FUNCTION "LKinLang_TokenizeSlot" : DWord   // FC35483, SCL
TITLE = LKinLang_TokenizeSlot
{ S7_Optimized_Access := 'TRUE' }
AUTHOR : tech.team.motioncontrol@siemens.com
FAMILY : LKinLang
VERSION : 1.1
// The FC separates a slot / line from line buffer in separate tokens
   VAR_INPUT
      lineNumber : UDInt;   // Line number input
      line : String;   // Line content input
      lastIndexOfMerger : Int;   // Last index of merger array
   END_VAR
   VAR_OUTPUT
      tokenizedLine : "LKinLang_typeLineTokens";   // Result of tokenization
   END_VAR
   VAR_IN_OUT
      separators : Array[1.."LKINLANG_NUMBER_OF_SEPARATORS"] of Byte;   // Array of separators
      mergers : Array[1.."LKINLANG_NUMBER_OF_MERGERS"] of Byte;   // Array of mergers
      preprocessorConfig : "LKinLang_typePreProcessorReplacement";   // Configuration structure for preProcessor (search/replace)
      errorString : String;   // Error in string format
   END_VAR
   VAR_TEMP
      tempAsciiLine : String["LKINLANG_LENGTH_OF_ASCII_LINE_STRING"];   // Temporary variable for the string line
      tempSeparatorIndex : DInt;   // Temporary variable for found separator index
      tempAsciiLineLength : Int;   // Temporary variable for the length of the string
      tempSignIndex : Int;   // Temporary counter in the string
      tempSignIndexOld : Int;   // Temporary old value of the counter in the string
      tempTokenIndex : Int;   // Temporary token counter for one line
      tempTypeOfChar : Array[0.."LKINLANG_LENGTH_OF_ASCII_LINE_STRING"] of USInt;   // Type of char in string: 0 = Defauflt; 1=Letter, 2=Number, 3=Merger
      tempTokenizedSlotEmpty : "LKinLang_typeLineTokens";   // Empty structure to delete last result
   END_VAR
   // Ret_Val : Return value of function
   VAR CONSTANT
      ERR_INVALID_LINE_NUMBER : DWord := 16#8200;   // Error due to wrong line number
      ERR_TOKEN_OVERFLOW : DWord := 16#8201;   // Error due to token being too long
      ERR_LINE_TOKEN_OUT_OF_BOUNDS : DWord := 16#8202;   // Error due to counter out of array bounds
   END_VAR
BEGIN
   //==========================================================================================
   // SIEMENS AG
   // (c)Copyright 2019 All Rights Reserved
   //------------------------------------------------------------------------------------------
   // Library: LKinLang
   // Tested with: S7-1517T-3 PN/DP
   // Engineering: TIA Portal V15
   // Restrictions: ---
   // Requirements: S7-1500T FW 2.5
   // Functionality: LKinLang_TokenizeSlot
   // The FC separates a slot / line from line buffer in separate tokens
   // 
   // Support: tech.team.motioncontrol@siemens.com
   // Note: Parameter comments are only available in language 'English (United States)'
   //------------------------------------------------------------------------------------------
   // Change log table:
   // Version    Date          Expert in charge    Changes applied
   // 01.00.00   28.05.2019    FR                  First created version
   // 02.00.00   20.03.2020    FR                  Changed funtion to work with one line only
   //=============================================================================

   // Intitialize values
   #LKinLang_TokenizeSlot := 0;
   #tempTokenIndex := 1;

   //--------------------------------------------------------------------------
   // All lines of Slot (PROGRAM) 
   // Information string access: first character to last character [1..n]
   // In Version 1.0 only one line of Slot (tempLineIndexMin == tempLineIndexMax)
   //--------------------------------------------------------------------------
   // FOR #tempLineIndex := #tempLineIndexMin TO #tempLineIndexMax DO

     // Init tokenized slot 
   #tokenizedLine := #tempTokenizedSlotEmpty;

     // Local copy OF ascii line
     #tempAsciiLine := #line;

     // Call of Pre Processor replacements
     "LKinLang_PreProcessor"(preprocessorConfig := #preprocessorConfig,
                             programLine := #tempAsciiLine);

     // Line which includes only a comment counts as an empty codeline (no G command)        
     "LKinLang_DeleteComment"(#tempAsciiLine);

     // Replace $T through space
     "LKinLang_ReplaceTapsBySpaces"(#tempAsciiLine);

     // Delete more than one spaces
     "LKinLang_DeleteMoreThanOneSpaceInRow"(#tempAsciiLine);

     // Length of ascii line
     #tempAsciiLineLength := LEN(#tempAsciiLine);

     IF #tempAsciiLineLength > 0 THEN
       // Get Tyoe of character --> write into array of USINT
       // Later check only Array and do not use Functions
       FOR #tempSignIndex := 1 TO #tempAsciiLineLength DO
         IF "LKinLang_CharacterIsLetter"(CHAR_TO_BYTE(#tempAsciiLine[#tempSignIndex])) THEN
           #tempTypeOfChar[#tempSignIndex] := 1;
         ELSIF "LKinLang_CharacterIsNumeric"(#tempAsciiLine[#tempSignIndex]) THEN
           #tempTypeOfChar[#tempSignIndex] := 2;
         ELSIF "LKinLang_CharacterIsMerger"(character := #tempAsciiLine[#tempSignIndex], lastIndexOfMerger := #lastIndexOfMerger, mergers := #mergers) THEN
           #tempTypeOfChar[#tempSignIndex] := 3;
         ELSE
           #tempTypeOfChar[#tempSignIndex] := 0;
         END_IF;
       END_FOR;

       #tempSignIndexOld := #tempAsciiLineLength + 1;

       // all characters of line
       FOR #tempSignIndex := #tempAsciiLineLength TO 1 BY -1 DO

         IF #tempTypeOfChar[#tempSignIndex] = 0 THEN // Only check for separator if not merger or letter or numeric: FR 2019.03.13
           REGION CECK_FOR_SEPARATOR
             //Check for separator
             //--------------------------------------------------------------------------------
             // compare sign with all separators
             FOR #tempSeparatorIndex := 1 TO "LKINLANG_NUMBER_OF_SEPARATORS" DO
               // detect separator
               IF #separators[#tempSeparatorIndex] = #tempAsciiLine[#tempSignIndex] THEN
                 IF #tempAsciiLineLength - #tempSignIndex > 0
                   AND #tempSignIndexOld - (#tempSignIndex + 1) > 0
                 THEN
                   IF #tempSignIndexOld - (#tempSignIndex + 1) <= "LKINLANG_LENGTH_OF_TOKEN_STRING" THEN
                     IF #tempTokenIndex > "LKINLANG_MAX_NUMBER_OF_TOKEN_PER_LINE" THEN
                       ;//Error: Array out of bounds 
                       #LKinLang_TokenizeSlot := #ERR_LINE_TOKEN_OUT_OF_BOUNDS;
                       #errorString := CONCAT(IN1 := #errorString, IN2 := 'Error: Tokenization - Overflow. Increase number of token per line - line: ');
                       #errorString := CONCAT(IN1 := #errorString, IN2 := UDINT_TO_STRING(#lineNumber));
                       RETURN;
                     ELSE
                       #tokenizedLine.lineToken[#tempTokenIndex] := MID(IN := #tempAsciiLine, P := #tempSignIndex + 1, L := #tempSignIndexOld - (#tempSignIndex + 1));
                       #tempTokenIndex := #tempTokenIndex + 1;
                     END_IF;
                   ELSE
                     ; // ERROR: Token overflow
                     #LKinLang_TokenizeSlot := #ERR_TOKEN_OVERFLOW;
                     #errorString := CONCAT(IN1 := #errorString, IN2 := 'Error: Tokenization - Overflow. Increase token length - line: ');
                     #errorString := CONCAT(IN1 := #errorString, IN2 := UDINT_TO_STRING(#lineNumber));
                     RETURN;
                   END_IF;
                 END_IF;

                 IF #tempTokenIndex > "LKINLANG_MAX_NUMBER_OF_TOKEN_PER_LINE" THEN
                   ;//Error: Array out of bounds 
                   #LKinLang_TokenizeSlot := #ERR_LINE_TOKEN_OUT_OF_BOUNDS;
                   #errorString := CONCAT(IN1 := #errorString, IN2 := 'Error: Tokenization - Overflow. Increase number of token per line - line: ');
                   #errorString := CONCAT(IN1 := #errorString, IN2 := UDINT_TO_STRING(#lineNumber));
                   RETURN;
                 ELSE
                   #tokenizedLine.lineToken[#tempTokenIndex] := MID(IN := #tempAsciiLine, P := #tempSignIndex, L := 1);
                   #tempTokenIndex := #tempTokenIndex + 1;
                   #tempSignIndexOld := #tempSignIndex;
                 END_IF;
                 EXIT;
               ELSE
                 ;// no match
               END_IF;
             END_FOR;
           END_REGION
         END_IF;

         REGION CHECK_FOR_LETTER_NUMBER
           //--------------------------------------------------------------------------------
           // Separator: Letter -> Number or Number -> letter
           IF #tempSignIndex >= 2 THEN // only possible if it isn´t the last character
             // Changed FR 2019.03.11: Replaced FC call with array
             IF
               ((#tempTypeOfChar[#tempSignIndex] = 2 AND (#tempTypeOfChar[#tempSignIndex - 1] = 1 OR NOT (#tempTypeOfChar[#tempSignIndex - 1] = 2))) // Number -> Letter 
               OR (#tempTypeOfChar[#tempSignIndex] = 1 AND (#tempTypeOfChar[#tempSignIndex - 1] = 2 OR NOT (#tempTypeOfChar[#tempSignIndex - 1] = 1)))) // Letter -> Number
               AND NOT (#tempTypeOfChar[#tempSignIndex - 1] = 3) // Merger to not separate Tokens
             THEN
               // New token found
               IF (#tempSignIndexOld - #tempSignIndex) <= "LKINLANG_LENGTH_OF_TOKEN_STRING" THEN
                 IF #tempTokenIndex > "LKINLANG_MAX_NUMBER_OF_TOKEN_PER_LINE" THEN
                   ;//Error: Array out of bounds 
                   #LKinLang_TokenizeSlot := #ERR_LINE_TOKEN_OUT_OF_BOUNDS;
                   #errorString := CONCAT(IN1 := #errorString, IN2 := 'Error: Tokenization - Overflow. Increase number of token per line - line: ');
                   #errorString := CONCAT(IN1 := #errorString, IN2 := UDINT_TO_STRING(#lineNumber));
                   RETURN;
                 ELSE
                   #tokenizedLine.lineToken[#tempTokenIndex] := MID(IN := #tempAsciiLine, P := #tempSignIndex, L := #tempSignIndexOld - #tempSignIndex);
                   #tempTokenIndex := #tempTokenIndex + 1;
                   #tempSignIndexOld := #tempSignIndex;
                 END_IF;
               ELSE
                 // ERROR: Token overflow
                 #LKinLang_TokenizeSlot := #ERR_TOKEN_OVERFLOW;
                 #errorString := CONCAT(IN1 := #errorString, IN2 := 'Error: Tokenization - Overflow. Increase token length');
                 RETURN;
               END_IF;
             ELSE
               ; // No change in character type --> check next character
             END_IF;
           END_IF;
           //--------------------------------------------------------------------------------
         END_REGION
       END_FOR;

       // Write number of token to structure
       #tokenizedLine.numberOfToken := INT_TO_UINT(#tempTokenIndex);

       // Last few signs
       IF #tempTokenIndex > "LKINLANG_MAX_NUMBER_OF_TOKEN_PER_LINE" THEN
         ;//Error: Array out of bounds 
         #LKinLang_TokenizeSlot := #ERR_LINE_TOKEN_OUT_OF_BOUNDS;
         #errorString := CONCAT(IN1 := #errorString, IN2 := 'Error: Tokenization - Overflow. Increase number of token per line - line: ');
         #errorString := CONCAT(IN1 := #errorString, IN2 := UDINT_TO_STRING(#lineNumber));
         RETURN;
       ELSE
         #tokenizedLine.lineToken[#tempTokenIndex] := MID(IN := #tempAsciiLine, P := 1, L := #tempSignIndexOld - 1);
       END_IF;
       // set token index for next line
       #tempTokenIndex := 1;
       // Write line number of ASCII file for N
       #tokenizedLine.lineNo := #lineNumber;

     ELSE
       // Empty line 
       #tokenizedLine.numberOfToken := 0;
       #tokenizedLine.lineNo := #lineNumber;
     END_IF;

   // END_FOR; //END: All lines of Slot (PROGRAM)
END_FUNCTION

FUNCTION "LKinLang_UpdateModalData" : Void   // FC35484, SCL
TITLE = LKinLang_UpdateModalData
{ S7_Optimized_Access := 'TRUE' }
AUTHOR : tech.team.motioncontrol@siemens.com
FAMILY : LKinLang
VERSION : 1.1
// The FC updates only modal parameters in a given PathData element
   VAR_IN_OUT
      inputPathData : "LKinLang_typePathDataElement";   // input PathData element to be updated
      updatedPathData : "LKinLang_typePathDataElement";   // updated PathData element
   END_VAR
   VAR_TEMP
      tempCounter : Int;   // temporary counter / temporary counter for empty lines
   END_VAR
BEGIN
   //==========================================================================================
   // SIEMENS AG
   // (c)Copyright 2019 All Rights Reserved
   //------------------------------------------------------------------------------------------
   // Library: LKinLang
   // Tested with: S7-1517T-3 PN/DP
   // Engineering: TIA Portal V15
   // Restrictions: ---
   // Requirements: S7-1500T FW 2.5
   // Functionality: LKinLang_UpdateModalData
   // The FC updates only modal parameters in a given PathData element
   // 
   // Support: tech.team.motioncontrol@siemens.com
   // Note: Parameter comments are only available in language 'English (United States)'
   //------------------------------------------------------------------------------------------
   // Change log table:
   // Version    Date          Expert in charge    Changes applied
   // 01.00.00   28.05.2019    FR                  First created version
   // 01.00.02   29.07.2019    FR                  Removed max negative value condition from IFs
   //=============================================================================

   //======================================================================
   // Copy input to output where input is not default and priority is higher
   //======================================================================  


   REGION UPDATE_ALL
     // Check CmdType
     IF #inputPathData.priority.cmdType > #updatedPathData.priority.cmdType THEN
       #updatedPathData.pathDataElement.cmdType := #inputPathData.pathDataElement.cmdType;
       #updatedPathData.priority.cmdType := #inputPathData.priority.cmdType;
     END_IF;

     // Check Coordinates
     // Update Cartesian positions
     IF  #inputPathData.priority.cmdCoordinates.cartesianPosition.x > #updatedPathData.priority.cmdCoordinates.cartesianPosition.x THEN
       #updatedPathData.pathDataElement.cmdCoordinates.cartesianPosition.x := #inputPathData.pathDataElement.cmdCoordinates.cartesianPosition.x;
       #updatedPathData.priority.cmdCoordinates.cartesianPosition.x := #inputPathData.priority.cmdCoordinates.cartesianPosition.x;
     END_IF;
     IF  #inputPathData.priority.cmdCoordinates.cartesianPosition.y > #updatedPathData.priority.cmdCoordinates.cartesianPosition.y THEN
       #updatedPathData.pathDataElement.cmdCoordinates.cartesianPosition.y := #inputPathData.pathDataElement.cmdCoordinates.cartesianPosition.y;
       #updatedPathData.priority.cmdCoordinates.cartesianPosition.y := #inputPathData.priority.cmdCoordinates.cartesianPosition.y;
     END_IF;
     IF  #inputPathData.priority.cmdCoordinates.cartesianPosition.z > #updatedPathData.priority.cmdCoordinates.cartesianPosition.z THEN
       #updatedPathData.pathDataElement.cmdCoordinates.cartesianPosition.z := #inputPathData.pathDataElement.cmdCoordinates.cartesianPosition.z;
       #updatedPathData.priority.cmdCoordinates.cartesianPosition.z := #inputPathData.priority.cmdCoordinates.cartesianPosition.z;
     END_IF;
     IF #inputPathData.priority.cmdCoordinates.cartesianPosition.a > #updatedPathData.priority.cmdCoordinates.cartesianPosition.a THEN
       #updatedPathData.pathDataElement.cmdCoordinates.cartesianPosition.a := #inputPathData.pathDataElement.cmdCoordinates.cartesianPosition.a;
       #updatedPathData.priority.cmdCoordinates.cartesianPosition.a := #inputPathData.priority.cmdCoordinates.cartesianPosition.a;
     END_IF;

     // Check coord system
     IF #inputPathData.priority.cmdCoordinates.coordSystem > #updatedPathData.priority.cmdCoordinates.coordSystem THEN
       #updatedPathData.pathDataElement.cmdCoordinates.coordSystem := #inputPathData.pathDataElement.cmdCoordinates.coordSystem;
       #updatedPathData.priority.cmdCoordinates.coordSystem := #inputPathData.priority.cmdCoordinates.coordSystem;
     END_IF;

     // Check Parameter
     // Check buffer mode
     IF #inputPathData.priority.cmdParameters.bufferMode > #updatedPathData.priority.cmdParameters.bufferMode THEN
       #updatedPathData.pathDataElement.cmdParameters.bufferMode := #inputPathData.pathDataElement.cmdParameters.bufferMode;
       #updatedPathData.priority.cmdParameters.bufferMode := #inputPathData.priority.cmdParameters.bufferMode;
     END_IF;

     // Check dynamic adaption
     IF #inputPathData.priority.cmdParameters.dynamicAdaption > #updatedPathData.priority.cmdParameters.dynamicAdaption THEN
       #updatedPathData.pathDataElement.cmdParameters.dynamicAdaption := #inputPathData.pathDataElement.cmdParameters.dynamicAdaption;
       #updatedPathData.priority.cmdParameters.dynamicAdaption := #inputPathData.priority.cmdParameters.dynamicAdaption;
     END_IF;

     // Check offsetParaNo
     IF #inputPathData.priority.cmdParameters.offsetParameters.offsetParaNo > #updatedPathData.priority.cmdParameters.offsetParameters.offsetParaNo THEN
       #updatedPathData.pathDataElement.cmdParameters.offsetParameters.offsetParaNo := #inputPathData.pathDataElement.cmdParameters.offsetParameters.offsetParaNo;
       #updatedPathData.priority.cmdParameters.offsetParameters.offsetParaNo := #inputPathData.priority.cmdParameters.offsetParameters.offsetParaNo;
     END_IF;

     // Check main path plane
     IF #inputPathData.priority.cmdParameters.offsetParameters.mainPathPlane > #updatedPathData.priority.cmdParameters.offsetParameters.mainPathPlane THEN
       #updatedPathData.pathDataElement.cmdParameters.offsetParameters.mainPathPlane := #inputPathData.pathDataElement.cmdParameters.offsetParameters.mainPathPlane;
       #updatedPathData.priority.cmdParameters.offsetParameters.mainPathPlane := #inputPathData.priority.cmdParameters.offsetParameters.mainPathPlane;
     END_IF;

     // Check orientation direction
     IF #inputPathData.priority.cmdParameters.orientationDirection > #updatedPathData.priority.cmdParameters.orientationDirection THEN
       #updatedPathData.pathDataElement.cmdParameters.orientationDirection := #inputPathData.pathDataElement.cmdParameters.orientationDirection;
       #updatedPathData.priority.cmdParameters.orientationDirection := #inputPathData.priority.cmdParameters.orientationDirection;
     END_IF;

     // Check transition parameter
     FOR #tempCounter := 1 TO 5 DO
       IF #inputPathData.priority.cmdParameters.transitionParameters[#tempCounter] > #updatedPathData.priority.cmdParameters.transitionParameters[#tempCounter] THEN
         #updatedPathData.pathDataElement.cmdParameters.transitionParameters[#tempCounter] := #inputPathData.pathDataElement.cmdParameters.transitionParameters[#tempCounter];
         #updatedPathData.priority.cmdParameters.transitionParameters[#tempCounter] := #inputPathData.priority.cmdParameters.transitionParameters[#tempCounter];
       END_IF;
     END_FOR;

     // Check circle parameters
     // Arc
     IF #inputPathData.priority.cmdParameters.circleParameters.arc > #updatedPathData.priority.cmdParameters.circleParameters.arc THEN
       #updatedPathData.pathDataElement.cmdParameters.circleParameters.arc := #inputPathData.pathDataElement.cmdParameters.circleParameters.arc;
       #updatedPathData.priority.cmdParameters.circleParameters.arc := #inputPathData.priority.cmdParameters.circleParameters.arc;
     END_IF;

     // Circ plane
     IF #inputPathData.priority.cmdParameters.circleParameters.circlePlane > #updatedPathData.priority.cmdParameters.circleParameters.circlePlane THEN
       #updatedPathData.pathDataElement.cmdParameters.circleParameters.circlePlane := #inputPathData.pathDataElement.cmdParameters.circleParameters.circlePlane;
       #updatedPathData.priority.cmdParameters.circleParameters.circlePlane := #inputPathData.priority.cmdParameters.circleParameters.circlePlane;
     END_IF;

     // Circ mode
     IF #inputPathData.priority.cmdParameters.circleParameters.circMode > #updatedPathData.priority.cmdParameters.circleParameters.circMode THEN
       #updatedPathData.pathDataElement.cmdParameters.circleParameters.circMode := #inputPathData.pathDataElement.cmdParameters.circleParameters.circMode;
       #updatedPathData.priority.cmdParameters.circleParameters.circMode := #inputPathData.priority.cmdParameters.circleParameters.circMode;
     END_IF;

     // path choice 
     IF #inputPathData.priority.cmdParameters.circleParameters.pathChoice > #updatedPathData.priority.cmdParameters.circleParameters.pathChoice THEN
       #updatedPathData.pathDataElement.cmdParameters.circleParameters.pathChoice := #inputPathData.pathDataElement.cmdParameters.circleParameters.pathChoice;
       #updatedPathData.priority.cmdParameters.circleParameters.pathChoice := #inputPathData.priority.cmdParameters.circleParameters.pathChoice;
     END_IF;

     // Radius
     IF #inputPathData.priority.cmdParameters.circleParameters.radius > #updatedPathData.priority.cmdParameters.circleParameters.radius THEN
       #updatedPathData.pathDataElement.cmdParameters.circleParameters.radius := #inputPathData.pathDataElement.cmdParameters.circleParameters.radius;
       #updatedPathData.priority.cmdParameters.circleParameters.radius := #inputPathData.priority.cmdParameters.circleParameters.radius;
     END_IF;

     // Aux point
     FOR #tempCounter := 1 TO 3 DO
       IF #inputPathData.priority.cmdParameters.circleParameters.auxPoint[#tempCounter] > #updatedPathData.priority.cmdParameters.circleParameters.auxPoint[#tempCounter] THEN
         #updatedPathData.pathDataElement.cmdParameters.circleParameters.auxPoint[#tempCounter] := #inputPathData.pathDataElement.cmdParameters.circleParameters.auxPoint[#tempCounter];
         #updatedPathData.priority.cmdParameters.circleParameters.auxPoint[#tempCounter] := #inputPathData.priority.cmdParameters.circleParameters.auxPoint[#tempCounter];
       END_IF;
     END_FOR;


     // Check dynamics
     // Velocity
     IF #inputPathData.priority.cmdParameters.pathDynamics.velocity > #updatedPathData.priority.cmdParameters.pathDynamics.velocity THEN
       #updatedPathData.pathDataElement.cmdParameters.pathDynamics.velocity := #inputPathData.pathDataElement.cmdParameters.pathDynamics.velocity;
       #updatedPathData.priority.cmdParameters.pathDynamics.velocity := #inputPathData.priority.cmdParameters.pathDynamics.velocity;
     END_IF;

     // Accelerration
     IF #inputPathData.priority.cmdParameters.pathDynamics.acceleration > #updatedPathData.priority.cmdParameters.pathDynamics.acceleration THEN
       #updatedPathData.pathDataElement.cmdParameters.pathDynamics.acceleration := #inputPathData.pathDataElement.cmdParameters.pathDynamics.acceleration;
       #updatedPathData.priority.cmdParameters.pathDynamics.acceleration := #inputPathData.priority.cmdParameters.pathDynamics.acceleration;
     END_IF;

     // Deceleration
     IF #inputPathData.priority.cmdParameters.pathDynamics.deceleration > #updatedPathData.priority.cmdParameters.pathDynamics.deceleration THEN
       #updatedPathData.pathDataElement.cmdParameters.pathDynamics.deceleration := #inputPathData.pathDataElement.cmdParameters.pathDynamics.deceleration;
       #updatedPathData.priority.cmdParameters.pathDynamics.deceleration := #inputPathData.priority.cmdParameters.pathDynamics.deceleration;
     END_IF;

     // Jerk
     IF #inputPathData.priority.cmdParameters.pathDynamics.jerk > #updatedPathData.priority.cmdParameters.pathDynamics.jerk THEN
       #updatedPathData.pathDataElement.cmdParameters.pathDynamics.jerk := #inputPathData.pathDataElement.cmdParameters.pathDynamics.jerk;
       #updatedPathData.priority.cmdParameters.pathDynamics.jerk := #inputPathData.priority.cmdParameters.pathDynamics.jerk;
     END_IF;

     // Check flags
     FOR #tempCounter := 1 TO "LKINCTRL_NO_OF_CMD_SETFLAGS" DO
       // Check set flag
       IF #inputPathData.priority.setFlags[#tempCounter].flag > #updatedPathData.priority.setFlags[#tempCounter].flag THEN
         #updatedPathData.pathDataElement.setFlags[#tempCounter].flag := #inputPathData.pathDataElement.setFlags[#tempCounter].flag;
         #updatedPathData.priority.setFlags[#tempCounter].flag := #inputPathData.priority.setFlags[#tempCounter].flag;
       END_IF;

       // Check flag mode
       IF #inputPathData.priority.setFlags[#tempCounter].flagMode > #updatedPathData.priority.setFlags[#tempCounter].flagMode THEN
         #updatedPathData.pathDataElement.setFlags[#tempCounter].flagMode := #inputPathData.pathDataElement.setFlags[#tempCounter].flagMode;
         #updatedPathData.priority.setFlags[#tempCounter].flagMode := #inputPathData.priority.setFlags[#tempCounter].flagMode;
       END_IF;

       // Check flag remaining distance
       IF #inputPathData.priority.setFlags[#tempCounter].flagMode > #updatedPathData.priority.setFlags[#tempCounter].remainingDistance THEN
         #updatedPathData.pathDataElement.setFlags[#tempCounter].remainingDistance := #inputPathData.pathDataElement.setFlags[#tempCounter].remainingDistance;
         #updatedPathData.priority.setFlags[#tempCounter].remainingDistance := #inputPathData.priority.setFlags[#tempCounter].remainingDistance;
       END_IF;
     END_FOR;

     // Check value flags
     FOR #tempCounter := 1 TO "LKINCTRL_NO_OF_CMD_VALUEFLAGS" DO
       // Check set flag
       IF #inputPathData.priority.valueFlags[#tempCounter].flag > #updatedPathData.priority.valueFlags[#tempCounter].flag THEN
         #updatedPathData.pathDataElement.valueFlags[#tempCounter].flag := #inputPathData.pathDataElement.valueFlags[#tempCounter].flag;
         #updatedPathData.priority.valueFlags[#tempCounter].flag := #inputPathData.priority.valueFlags[#tempCounter].flag;
       END_IF;

       // Check flag mode
       IF #inputPathData.priority.valueFlags[#tempCounter].flagMode > #updatedPathData.priority.valueFlags[#tempCounter].flagMode THEN
         #updatedPathData.pathDataElement.valueFlags[#tempCounter].flagMode := #inputPathData.pathDataElement.valueFlags[#tempCounter].flagMode;
         #updatedPathData.priority.valueFlags[#tempCounter].flagMode := #inputPathData.priority.valueFlags[#tempCounter].flagMode;
       END_IF;

       // Check flag remaining distance
       IF #inputPathData.priority.valueFlags[#tempCounter].flagMode > #updatedPathData.priority.valueFlags[#tempCounter].remainingDistance THEN
         #updatedPathData.pathDataElement.valueFlags[#tempCounter].remainingDistance := #inputPathData.pathDataElement.valueFlags[#tempCounter].remainingDistance;
         #updatedPathData.priority.valueFlags[#tempCounter].remainingDistance := #inputPathData.priority.valueFlags[#tempCounter].remainingDistance;
       END_IF;
     END_FOR;
   END_REGION
END_FUNCTION

FUNCTION "LKinLang_GetVariable" : Void   // FC35485, SCL
TITLE = LKinLang_GetVariable
{ S7_Optimized_Access := 'TRUE' }
AUTHOR : tech.team.motioncontrol@siemens.com
FAMILY : LKinLang
VERSION : 1.0
// The FC gets the value of a variable and adds it to a string
   VAR_INPUT
      varIndex : Int;   // Variable index
      varType : Int;   // Variable type
   END_VAR
   VAR_IN_OUT
      localVariables : "LKinLang_typeLocalVariables";   // Variables reference list
      interfaceVariables : "LKinLang_typeInterfaceVariables";   // Key token to find variables
      stringExpression : String;   // String expression
   END_VAR
BEGIN
   //==========================================================================================
   // SIEMENS AG
   // (c)Copyright 2020 All Rights Reserved
   //------------------------------------------------------------------------------------------
   // Library: LKinLang
   // Tested with: S7-1517T-3 PN/DP
   // Engineering: TIA Portal V15
   // Restrictions: ---
   // Requirements: S7-1500T FW 2.5
   // Functionality: LKinLang_IsTokenVariable
   // The FC gets the value of a variable and adds it to a string
   // 
   // Support: tech.team.motioncontrol@siemens.com
   // Note: Parameter comments are only available in language 'English (United States)'
   //------------------------------------------------------------------------------------------
   // Change log table:
   // Version    Date          Expert in charge    Changes applied
   // 01.00.00   24.11.2020    FR                  First created version
   //===========================================================================================

   // --------------------------------------------------------------
   // Right side of equation 
   // --> GET value of variable
   // Concat to string expression
   // --------------------------------------------------------------
   CASE #varType OF
     "LKINLANG_VAR_TYPE_LOCAL_BOOL": // local bool
       // Concat value of var to string expression    
       #stringExpression := CONCAT(IN1 := DINT_TO_STRING(BOOL_TO_DINT(#localVariables.boolean[#varIndex])),
                                       IN2 := #stringExpression);

       // 16.07.2019 FR: Delete "+" sign from string
       IF BOOL_TO_DINT(#localVariables.boolean[#varIndex]) >= 0.0 THEN
         #stringExpression := DELETE(IN := #stringExpression, L := 1, P := 1);
       ELSE
         ; // Keep "-" sign
       END_IF;


     "LKINLANG_VAR_TYPE_LOCAL_DINT": // local dint
       // Concat value of var to string expression    
       #stringExpression := CONCAT(IN1 := DINT_TO_STRING(#localVariables.dints[#varIndex]),
                                       IN2 := #stringExpression);

       // 16.07.2019 FR: Delete "+" sign from string
       IF #localVariables.dints[#varIndex] >= 0.0 THEN
         #stringExpression := DELETE(IN := #stringExpression, L := 1, P := 1);
       ELSE
         ; // Keep "-" sign
       END_IF;

     "LKINLANG_VAR_TYPE_LOCAL_LREAL": // local lreal
       // Concat value of var to string expression
       #stringExpression := CONCAT(IN1 := "LKinLang_LRealToReducedString"(input := #localVariables.lreals[#varIndex], decimalPlaces := 6),
                                       IN2 := #stringExpression);


     "LKINLANG_VAR_TYPE_INTERFACE_BOOL":
       // Concat value of var to string expression    
       #stringExpression := CONCAT(IN1 := DINT_TO_STRING(BOOL_TO_DINT(#interfaceVariables.Boolean[#varIndex])),
                                       IN2 := #stringExpression);

       // 16.07.2019 FR: Delete "+" sign from string
       IF BOOL_TO_DINT(#interfaceVariables.Boolean[#varIndex]) >= 0.0 THEN
         #stringExpression := DELETE(IN := #stringExpression, L := 1, P := 1);
       ELSE
         ; // Keep "-" sign
       END_IF;

     "LKINLANG_VAR_TYPE_INTERFACE_DINT":
       // Get value of interface variable at given index
       // Concat value of var to string expression    
       #stringExpression := CONCAT(IN1 := DINT_TO_STRING(#interfaceVariables.DInts[#varIndex]),
                                       IN2 := #stringExpression);

       // Delete "+" sign from string
       IF #interfaceVariables.DInts[#varIndex] >= 0.0 THEN
         #stringExpression := DELETE(IN := #stringExpression, L := 1, P := 1);
       ELSE
         ; // Keep "-" sign
       END_IF;


     "LKINLANG_VAR_TYPE_INTERFACE_LREAL":
       // Concat value of var to string expression
       #stringExpression := CONCAT(IN1 := "LKinLang_LRealToReducedString"(input := #interfaceVariables.LReals[#varIndex], decimalPlaces := 6),
                                       IN2 := #stringExpression);

     ELSE
       ; // type not defined
   END_CASE;
END_FUNCTION

FUNCTION "LKinLang_SetVariable" : Void   // FC35486, SCL
TITLE = LKinLang_SetVariable
{ S7_Optimized_Access := 'TRUE' }
AUTHOR : tech.team.motioncontrol@siemens.com
FAMILY : LKinLang
VERSION : 1.0
// The FC checks a string for a value and sets the variable accordingly
   VAR_INPUT
      varIndex : Int;   // Variable index
      varType : Int;   // Variable type
      lineNumber : UDInt;   // Line number
   END_VAR
   VAR_IN_OUT
      stringExpression : String;   // String expression
      localVariables : "LKinLang_typeLocalVariables";   // Variables reference list
      interfaceVariables : "LKinLang_typeInterfaceVariables";   // Key token to find variables
      errorString : String;   // Error string connection
   END_VAR
   VAR_TEMP
      tempCounter : DInt;   // Temporary counter
      tempParameterValue : LReal;   // Temporary parameter value
      tempMathParserResult : "LKinLang_typeMathParserResult";   // Temporary result of math parser
   END_VAR
   VAR CONSTANT
      MINVAL_DINT : DInt := -2147483648 ;   // Minimum value of DINT
      MAXVAL_DINT : DInt := +2147483647;   // Minimum value of DINT
   END_VAR
BEGIN
   //==========================================================================================
   // SIEMENS AG
   // (c)Copyright 2020 All Rights Reserved
   //------------------------------------------------------------------------------------------
   // Library: LKinLang
   // Tested with: S7-1517T-3 PN/DP
   // Engineering: TIA Portal V15
   // Restrictions: ---
   // Requirements: S7-1500T FW 2.5
   // Functionality: LKinLang_IsTokenVariable
   // The FC checks a string for a value and sets the variable accordingly
   // 
   // Support: tech.team.motioncontrol@siemens.com
   // Note: Parameter comments are only available in language 'English (United States)'
   //------------------------------------------------------------------------------------------
   // Change log table:
   // Version    Date          Expert in charge    Changes applied
   // 01.00.00   24.11.2020    FR                  First created version
   //===========================================================================================

   // Check for TRUE in stringExpression
   #tempCounter := FIND(IN1 := #stringExpression, IN2 := 'TRUE');

   // Check if string expression contains TRUE / FALSE
   IF #tempCounter <> 0 AND (#varType = "LKINLANG_VAR_TYPE_INTERFACE_BOOL" OR #varType = "LKINLANG_VAR_TYPE_LOCAL_BOOL") THEN
     #stringExpression := REPLACE(IN1 := #stringExpression, IN2 := '1', L := 4, P := #tempCounter);
   ELSIF #tempCounter <> 0 AND (#varType <> "LKINLANG_VAR_TYPE_INTERFACE_BOOL" AND #varType <> "LKINLANG_VAR_TYPE_LOCAL_BOOL") THEN
     ;// Error using "TRUE" for wrong data type
     #errorString := CONCAT(IN1 := #errorString, IN2 := ';Error: No implicit dataType conversion possible');
     #errorString := CONCAT(IN1 := #errorString, IN2 := ' in line: ');
     #errorString := CONCAT(IN1 := #errorString, IN2 := UDINT_TO_STRING(#lineNumber));
   END_IF;

   // Check for FALSE in stringExpression
   #tempCounter := FIND(IN1 := #stringExpression, IN2 := 'FALSE');

   // Check if string expression contains TRUE / FALSE
   IF #tempCounter <> 0 AND (#varType = "LKINLANG_VAR_TYPE_INTERFACE_BOOL" OR #varType = "LKINLANG_VAR_TYPE_LOCAL_BOOL") THEN
     #stringExpression := REPLACE(IN1 := #stringExpression, IN2 := '0', L := 5, P := #tempCounter);
   ELSIF #tempCounter <> 0 AND (#varType <> "LKINLANG_VAR_TYPE_INTERFACE_BOOL" AND #varType <> "LKINLANG_VAR_TYPE_LOCAL_BOOL") THEN
     ;// Error using "FALSE" for wrong data type
     #errorString := CONCAT(IN1 := #errorString, IN2 := ';Error: No implicit dataType conversion possible');
     #errorString := CONCAT(IN1 := #errorString, IN2 := ' in line: ');
     #errorString := CONCAT(IN1 := #errorString, IN2 := UDINT_TO_STRING(#lineNumber));
   END_IF;

   // Check if string expression is just a number
   IF "LKinLang_IsTokenNumberInclSign"(#stringExpression) THEN
     // If just a number then directly assign value
     #tempParameterValue := STRING_TO_LREAL(#stringExpression);
   ELSE
     // Not a single number --> Use mathParser to calculate value
     #tempMathParserResult := "LKinLang_CalcMathAndBool"(inputString := #stringExpression);

     // Check for error in math parser
     IF #tempMathParserResult.errorID <> 0 THEN
       #errorString := CONCAT(IN1 := #errorString, IN2 := ';Error: Stringexpression ');
       #errorString := CONCAT(IN1 := #errorString, IN2 := #stringExpression);
     ELSE
       // Math parser delivers a valid result
       // Assign result to value
       #tempParameterValue := #tempMathParserResult.finalResult;
     END_IF;
   END_IF;

   // Set variable depending on type
   // Check if value fits into dataType
   CASE #varType OF
     "LKINLANG_VAR_TYPE_LOCAL_BOOL": // local bool
       IF #tempParameterValue <> 0.0 AND #tempParameterValue <> 1.0 THEN
         // Error variable overflow
         #errorString := CONCAT(IN1 := #errorString, IN2 := ';Error: Value exceeds size of local bool variable in line ');
         #errorString := CONCAT(IN1 := #errorString, IN2 := UDINT_TO_STRING(#lineNumber));
       ELSE
         #localVariables.boolean[#varIndex] := (#tempParameterValue = 1.0); // If 1.0 then true else false
       END_IF;

     "LKINLANG_VAR_TYPE_LOCAL_DINT": // local dint
       IF #tempParameterValue > #MAXVAL_DINT OR #tempParameterValue < #MINVAL_DINT THEN
         // Error variable overflow
         #errorString := CONCAT(IN1 := #errorString, IN2 := ';Error: Value exceeds size of local DInt variable in line ');
         #errorString := CONCAT(IN1 := #errorString, IN2 := UDINT_TO_STRING(#lineNumber));

       ELSE
         // Assing value
         #localVariables.dints[#varIndex] := LREAL_TO_DINT(#tempParameterValue);
       END_IF;

     "LKINLANG_VAR_TYPE_LOCAL_LREAL": // local lreal
       #localVariables.lreals[#varIndex] := #tempParameterValue;

     "LKINLANG_VAR_TYPE_INTERFACE_BOOL": // Interface bool
       IF #tempParameterValue <> 0.0 AND #tempParameterValue <> 1.0 THEN
         // Error variable overflow
         #errorString := CONCAT(IN1 := #errorString, IN2 := ';Error: Value exceeds size of Bool interface variable in line ');
         #errorString := CONCAT(IN1 := #errorString, IN2 := UDINT_TO_STRING(#lineNumber));
       ELSE
         #interfaceVariables.Boolean[#varIndex] := (#tempParameterValue = 1.0); // If 1.0 then true else false
       END_IF;

     "LKINLANG_VAR_TYPE_INTERFACE_DINT": // interface dint
       IF #tempParameterValue > #MAXVAL_DINT OR #tempParameterValue < #MINVAL_DINT THEN
         // Error variable overflow
         #errorString := CONCAT(IN1 := #errorString, IN2 := ';Error: Value exceeds size of DInt interface variable in line ');
         #errorString := CONCAT(IN1 := #errorString, IN2 := UDINT_TO_STRING(#lineNumber));
       ELSE
         #interfaceVariables.DInts[#varIndex] := LREAL_TO_DINT(#tempParameterValue);
       END_IF;

     "LKINLANG_VAR_TYPE_INTERFACE_LREAL": // interface lreal
       #interfaceVariables.LReals[#varIndex] := #tempParameterValue;

     ELSE
       ; // type not defined
   END_CASE;
END_FUNCTION

FUNCTION "LKinLang_IsTokenKeyWord" : Bool   // FC35488, SCL
TITLE = LKinLang_IsTokenKey / LKinLang_IsTokenKeyWord
{ S7_Optimized_Access := 'TRUE' }
AUTHOR : tech.team.motioncontrol@siemens.com
FAMILY : LKinLang
VERSION : 1.0
// The FC checks if a given token is a keyword
   VAR_INPUT
      token : String;   // Token to be check
   END_VAR
   VAR_IN_OUT
      keyToken : "LKinLang_typeKeyToken";   // Key token list
   END_VAR
   // Ret_Val : TRUE: Token is keyword; FALSE: Token is not a keyword
BEGIN
   //==========================================================================================
   // SIEMENS AG
   // (c)Copyright 2020 All Rights Reserved
   //------------------------------------------------------------------------------------------
   // Library: LKinLang
   // Tested with: S7-1517T-3 PN/DP
   // Engineering: TIA Portal V15
   // Restrictions: ---
   // Requirements: S7-1500T FW 2.5
   // Functionality: LKinLang_IsTokenVariable
   // The FC checks if a given token is a keyword
   // 
   // Support: tech.team.motioncontrol@siemens.com
   // Note: Parameter comments are only available in language 'English (United States)'
   //------------------------------------------------------------------------------------------
   // Change log table:
   // Version    Date          Expert in charge    Changes applied
   // 01.00.00   24.11.2020    FR                  First created version
   //===========================================================================================

   //======================================================================
   // Is token (or any other string) a keyword
   //======================================================================
   IF #token = #keyToken.tokenBool
       OR #token = #keyToken.tokenDInt
       OR #token = #keyToken.tokenLReal
       OR #token = #keyToken.tokenInterfaceVarBool
       OR #token = #keyToken.tokenInterfaceVarDInt
       OR #token = #keyToken.tokenInterfaceVarLReal
       OR #token = #keyToken.tokenJumpTarget
       OR #token = #keyToken.tokenJump
       OR #token = #keyToken.tokenJumpConditional
       OR #token = #keyToken.tokenPreprocessingStop
       OR #token = #keyToken.tokenIf
       OR #token = #keyToken.tokenElse
       OR #token = #keyToken.tokenEndIf
       OR #token = #keyToken.tokenWhile
       OR #token = #keyToken.tokenEndWhile
       OR #token = #keyToken.tokenFor
       OR #token = #keyToken.tokenQuantity
       OR #token = #keyToken.tokenIncrement
       OR #token = #keyToken.tokenEndFor
       OR #token = #keyToken.tokenStartSub
       OR #token = #keyToken.tokenEndSub
       OR #token = #keyToken.tokenCallSub
   THEN
       #LKinLang_IsTokenKeyWord := TRUE;
   ELSE
       #LKinLang_IsTokenKeyWord := FALSE;
   END_IF;
END_FUNCTION

(* ===== HMI "HMI_RT_1" =====
system functions are stored by id; their names below are inferred from use
connection "HMI_Connection_1": ETHERNET, S7_1500_OMS

HMI tags "Default tag table"
   "AxesEnabled" : Bool = PLC DB_Writing.AxesEnabled AT %DB1.DBX0.0, 1 s
   "AxesError" : Bool = PLC DB_Writing.AxesError AT %DB1.DBX0.0, 1 s
   "AxesHomed" : Bool = PLC DB_Writing.AxesHomed AT %DB1.DBX0.0, 1 s
   "EnableAxes" : Bool = PLC DB_Writing.EnableAxes AT %DB1.DBX0.0, 1 s
   "executeProgram" : Bool = PLC DB_Writing.executeProgram AT %DB1.DBX0.0, 1 s
   "HomeAxes" : Bool = PLC DB_Writing.HomeAxes AT %DB1.DBX0.0, 1 s
   "movePath_active" : Bool = PLC DB_Writing.movePath_active AT %DB1.DBX0.0, 1 s
   "movePath_status" : Word = PLC DB_Writing.movePath_status AT %DB1.DBW0, 1 s
   "programStatusString" : String[254] = PLC DB_Writing.programStatusString AT %DB1.DBW0, 1 s
   "ResetAxes" : Bool = PLC DB_Writing.ResetAxes AT %DB1.DBX0.0, 1 s
   "resetProgram" : Bool = PLC DB_Writing.resetProgram AT %DB1.DBX0.0, 1 s
   "stopProgram" : Bool = PLC DB_Writing.stopProgram AT %DB1.DBX0.0, 1 s
   "text" : String[254] = PLC DB_Writing.textInput AT %DB1.DBW0, 1 s
   "triggerProcessText" : Bool = PLC DB_Writing.triggerTextbox AT %DB1.DBX0.0, 1 s

screen "Writing_controls" 800x480
   TextField "Txt_AxStatus_1" at 332,286 size 60x21; Text 'Homed'
   TextField "Txt_AxStatus_2" at 332,319 size 67x21; Text 'Enabled'
   TextField "Txt_AxStatus_3" at 332,352 size 46x21; Text 'Error'
   TextField "Txt_Step_1" at 21,38 size 175x23; Text '1. Write your text:'
   TextField "Txt_Step_3" at 332,38 size 150x23; Text '2. Control axes:'
   TextField "Txt_Step_4" at 580,38 size 184x23; Text '3. Control program:'
   TextField "Txt_Status_1" at 21,254 size 166x24; Text 'Kinematics status'
   TextField "Txt_Status_2" at 332,254 size 111x24; Text 'Axes status'
   TextField "Txt_Status_3" at 580,254 size 144x24; Text 'Program status'
   Circle "LED_Axes_1" at 414,286 size 21x21
      Appearance <- "AxesHomed"
   Circle "LED_Axes_2" at 414,319 size 21x21
      Appearance <- "AxesEnabled"
   Circle "LED_Axes_3" at 414,352 size 21x21
      Appearance <- "AxesError"
   IOField "ProgramStatus" at 518,286 size 280x32; FormatPattern ??????????????????????????????
      ProcessValue <- "programStatusString"
   IOField "Input_text_field" at 22,77 size 264x32; FormatPattern ????????????????????
      ProcessValue <- "text"
      on Activate: ResetBit("triggerProcessText")
      on OnFinishInput: SetBit("triggerProcessText")
   SymbolicIOField "KineStatus_1" at 22,290 size 174x32; TextOff '0'; TextOn '1'; TextList "TextList_MovePathStatus"
      ProcessValue <- "movePath_status"
   SymbolicIOField "KineStatus_2" at 22,339 size 174x32; TextOn 'Kinematics in motion'; TextOff 'Standstill'
      ProcessValue <- "movePath_active"
   Switch "Switch_ExecuteProgram" at 580,71 size 163x38; TextOn 'Execute program'; CaptionText 'Switch'; TextOff 'Execute program'
      ProcessValue <- "executeProgram"
      Appearance <- "executeProgram"
   Switch "Switch_EnableAxes" at 332,119 size 142x38; TextOn 'Disable axes'; CaptionText 'Switch'; TextOff 'Enable axes'
      ProcessValue <- "EnableAxes"
      Appearance <- "EnableAxes"
   Switch "Switch_ResetAxes" at 332,166 size 142x38; TextOn 'Reset axes'; CaptionText 'Switch'; TextOff 'Reset axes'
      ProcessValue <- "ResetAxes"
      Appearance <- "ResetAxes"
   Switch "Switch_HomeAxes" at 332,71 size 141x38; TextOn 'Home axes'; CaptionText 'Switch'; TextOff 'Home axes'
      ProcessValue <- "HomeAxes"
      Appearance <- "HomeAxes"
   Switch "Switch_StopProgram" at 580,119 size 163x38; TextOn 'Stop program'; CaptionText 'Switch'; TextOff 'Stop program'
      ProcessValue <- "stopProgram"
      Appearance <- "stopProgram"
   Switch "Switch_ResetProgram" at 580,166 size 163x38; TextOn 'Reset program'; CaptionText 'Switch'; TextOff 'Reset program'
      ProcessValue <- "resetProgram"
      Appearance <- "resetProgram"
*)